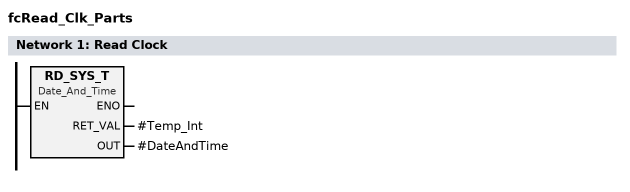
   #Temp_Int := RD_SYS_T(out => #DateAndTime);
END_REGION

REGION Network 2 (STL)

         LAR1  #""Address_4";
         L     B[AR1, P#0.0];
         T     #Year;
         L     B[AR1, P#1.0];
         T     #Month;
         L     B[AR1, P#2.0];
         T     #Day;
         L     B[AR1, P#3.0];
         T     #Hour;
         L     B[AR1, P#4.0];
         T     #Minute;
         L     B[AR1, P#5.0];
         T     #Second;

         L     W#16#FFF0;
         L     W[AR1, P#6.0];
         AW;
         T     #MilliSecond;

         L     B#16#F;
         L     B[AR1, P#7.0];
         AW;
         T     #DayOfWeek;
         CLR;
END_REGION
END_FUNCTION

FUNCTION "fcByteToBits" : Void   // FC1002, LAD
TITLE = Split byte into bits
{ S7_Optimized_Access := 'FALSE' }
VERSION : 0.1
BEGIN

REGION Network 1: Bit 0
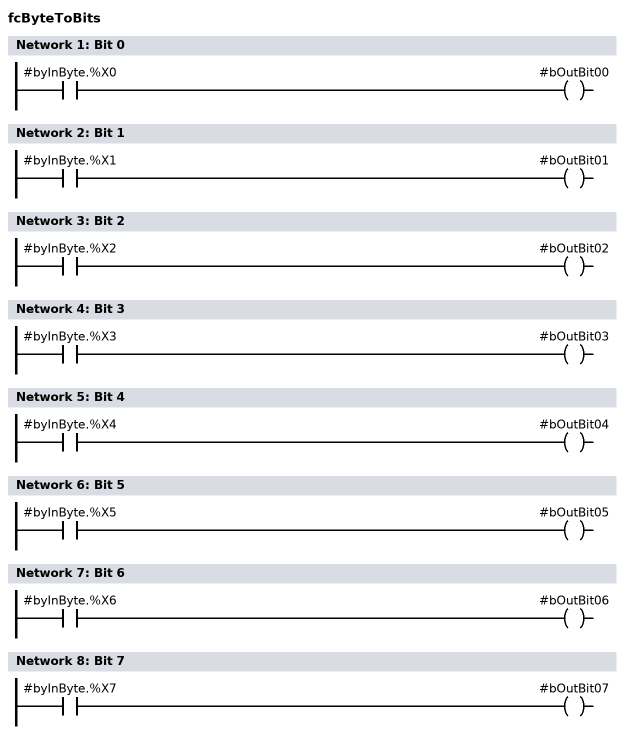
   RUNG wire#powerrail
      Contact( #byInByte.%X0 )
      Coil( #bOutBit00 )
   END_RUNG
   // the same network as SCL:
   #bOutBit00 := #byInByte.%X0;
END_REGION

REGION Network 2: Bit 1
   RUNG wire#powerrail
      Contact( #byInByte.%X1 )
      Coil( #bOutBit01 )
   END_RUNG
   // the same network as SCL:
   #bOutBit01 := #byInByte.%X1;
END_REGION

REGION Network 3: Bit 2
   RUNG wire#powerrail
      Contact( #byInByte.%X2 )
      Coil( #bOutBit02 )
   END_RUNG
   // the same network as SCL:
   #bOutBit02 := #byInByte.%X2;
END_REGION

REGION Network 4: Bit 3
   RUNG wire#powerrail
      Contact( #byInByte.%X3 )
      Coil( #bOutBit03 )
   END_RUNG
   // the same network as SCL:
   #bOutBit03 := #byInByte.%X3;
END_REGION

REGION Network 5: Bit 4
   RUNG wire#powerrail
      Contact( #byInByte.%X4 )
      Coil( #bOutBit04 )
   END_RUNG
   // the same network as SCL:
   #bOutBit04 := #byInByte.%X4;
END_REGION

REGION Network 6: Bit 5
   RUNG wire#powerrail
      Contact( #byInByte.%X5 )
      Coil( #bOutBit05 )
   END_RUNG
   // the same network as SCL:
   #bOutBit05 := #byInByte.%X5;
END_REGION

REGION Network 7: Bit 6
   RUNG wire#powerrail
      Contact( #byInByte.%X6 )
      Coil( #bOutBit06 )
   END_RUNG
   // the same network as SCL:
   #bOutBit06 := #byInByte.%X6;
END_REGION

REGION Network 8: Bit 7
   RUNG wire#powerrail
      Contact( #byInByte.%X7 )
      Coil( #bOutBit07 )
   END_RUNG
   // the same network as SCL:
   #bOutBit07 := #byInByte.%X7;
END_REGION
END_FUNCTION

FUNCTION "fbBitsToByte" : Void   // FC1003, LAD
TITLE = Pack bits into byte
{ S7_Optimized_Access := 'FALSE' }
VERSION : 0.1
BEGIN

REGION Network 1: Bit0
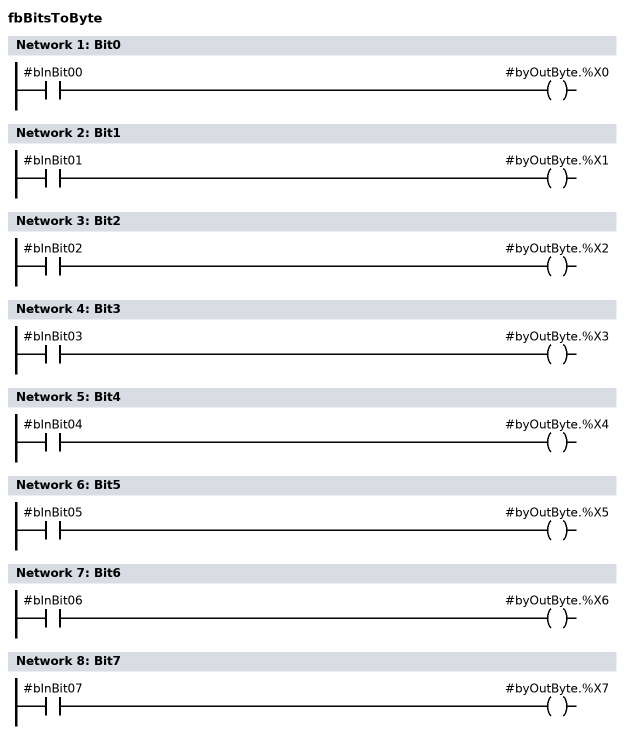
   RUNG wire#powerrail
      Contact( #bInBit00 )
      Coil( #byOutByte.%X0 )
   END_RUNG
   // the same network as SCL:
   #byOutByte.%X0 := #bInBit00;
END_REGION

REGION Network 2: Bit1
   RUNG wire#powerrail
      Contact( #bInBit01 )
      Coil( #byOutByte.%X1 )
   END_RUNG
   // the same network as SCL:
   #byOutByte.%X1 := #bInBit01;
END_REGION

REGION Network 3: Bit2
   RUNG wire#powerrail
      Contact( #bInBit02 )
      Coil( #byOutByte.%X2 )
   END_RUNG
   // the same network as SCL:
   #byOutByte.%X2 := #bInBit02;
END_REGION

REGION Network 4: Bit3
   RUNG wire#powerrail
      Contact( #bInBit03 )
      Coil( #byOutByte.%X3 )
   END_RUNG
   // the same network as SCL:
   #byOutByte.%X3 := #bInBit03;
END_REGION

REGION Network 5: Bit4
   RUNG wire#powerrail
      Contact( #bInBit04 )
      Coil( #byOutByte.%X4 )
   END_RUNG
   // the same network as SCL:
   #byOutByte.%X4 := #bInBit04;
END_REGION

REGION Network 6: Bit5
   RUNG wire#powerrail
      Contact( #bInBit05 )
      Coil( #byOutByte.%X5 )
   END_RUNG
   // the same network as SCL:
   #byOutByte.%X5 := #bInBit05;
END_REGION

REGION Network 7: Bit6
   RUNG wire#powerrail
      Contact( #bInBit06 )
      Coil( #byOutByte.%X6 )
   END_RUNG
   // the same network as SCL:
   #byOutByte.%X6 := #bInBit06;
END_REGION

REGION Network 8: Bit7
   RUNG wire#powerrail
      Contact( #bInBit07 )
      Coil( #byOutByte.%X7 )
   END_RUNG
   // the same network as SCL:
   #byOutByte.%X7 := #bInBit07;
END_REGION
END_FUNCTION

FUNCTION "fcCreateAnyPointer" : Void   // FC1025, STL
TITLE = Creates any pointer
{ S7_Optimized_Access := 'FALSE' }
VERSION : 0.1
BEGIN

REGION Network 1: It won't work in LAD, STL only
   // Create pointer in the temp location (AR1)
         LAR1  #""Address_2";

   // Syntax ID - always 10
         L     B#16#10;
         T     LB[AR1, P#0.0];

   // Data type
         L     #byInDataType;
         T     LB[AR1, P#1.0];

   // Size
         L     #iInSize;
         T     LW[AR1, P#2.0];

   // DB number
         L     #iInDB_Num;
         T     LW[AR1, P#4.0];


   // Memory area
         L     #byInMemoryArea;
         T     LB[AR1, P#6.0];

   // Offset high byte
         L     #iInOffsetByte;
         SRD   13;
         T     LB[AR1, P#7.0];

   // Offset low word
         L     #iInOffsetBit;
         AW    16#0007;

         L     #iInOffsetByte;
         SLD   3;

         OW;
         T     LW[AR1, P#8.0];

   // Write to the output (AR2)
         L     #""Address_21";
         LAR2;

         L     LD[AR1, P#0.0];
         T     D[AR2, P#0.0];

         L     LD[AR1, P#4.0];
         T     D[AR2, P#4.0];

         L     LW[AR1, P#8.0];
         T     W[AR2, P#8.0];
END_REGION

REGION Network 2
         SET;
         SAVE;
END_REGION
END_FUNCTION

FUNCTION "fcParseAnyPointer" : Void   // FC1026, SCL
{ S7_Optimized_Access := 'FALSE' }
VERSION : 0.0
BEGIN


       #AnyPointer := #pInAnyPointer;

       #AnyStruc.SyntaxID := b#16#10;
       #byOutDataType := #AnyStruc.DataType;
       #iOutSize := WORD_TO_INT(#AnyStruc.Size);
       #iOutDB_Num := WORD_TO_INT(#AnyStruc.DB_Num);
       #byOutMemoryArea := #AnyStruc.MemoryArea;
       #iOutOffsetBit := WORD_TO_INT(#AnyStruc.OffsetLo AND w#16#0007);
       #iOutOffsetByte := WORD_TO_INT(SHR(IN := #AnyStruc.OffsetLo, N := 3) OR SHL(IN := BYTE_TO_WORD(#AnyStruc.OffsetHi), N := 13));

       ENO:=true;
END_FUNCTION

FUNCTION "fcTemperatureConvert" : Void   // FC1027, LAD
{ S7_Optimized_Access := 'FALSE' }
VERSION : 0.1
BEGIN

REGION Network 1: Convert F to C
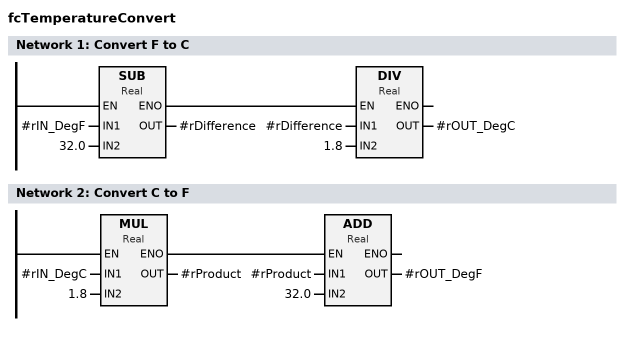
   RUNG wire#powerrail
      { S7_Templates := "SrcType := Real"; S7_GenerateENO := "TRUE" } Sub(in1 := #rIN_DegF, in2 := 32.0, out => #rDifference)
      { S7_Templates := "SrcType := Real"; S7_GenerateENO := "TRUE" } Div(in1 := #rDifference, in2 := 1.8, out => #rOUT_DegC)
   END_RUNG
   // the same network as SCL:
   // ENO of a box is taken as its EN; it also drops when the box reports an error
   #rDifference := #rIN_DegF - 32.0;
   #rOUT_DegC := #rDifference / 1.8;
END_REGION

REGION Network 2: Convert C to F
   RUNG wire#powerrail
      { S7_Templates := "SrcType := Real"; S7_GenerateENO := "TRUE" } Mul(in1 := #rIN_DegC, in2 := 1.8, out => #rProduct)
      { S7_Templates := "SrcType := Real"; S7_GenerateENO := "TRUE" } Add(in1 := #rProduct, in2 := 32.0, out => #rOUT_DegF)
   END_RUNG
   // the same network as SCL:
   // ENO of a box is taken as its EN; it also drops when the box reports an error
   #rProduct := #rIN_DegC * 1.8;
   #rOUT_DegF := #rProduct + 32.0;
END_REGION
END_FUNCTION

// folder: Resources/IO

FUNCTION "fcReadInput_LinearScale" : Void   // FC308, LAD
TITLE = Read/Scale input word
{ S7_Optimized_Access := 'FALSE' }
VERSION : 0.1
BEGIN

REGION Network 1: Swap input value bytes if needed
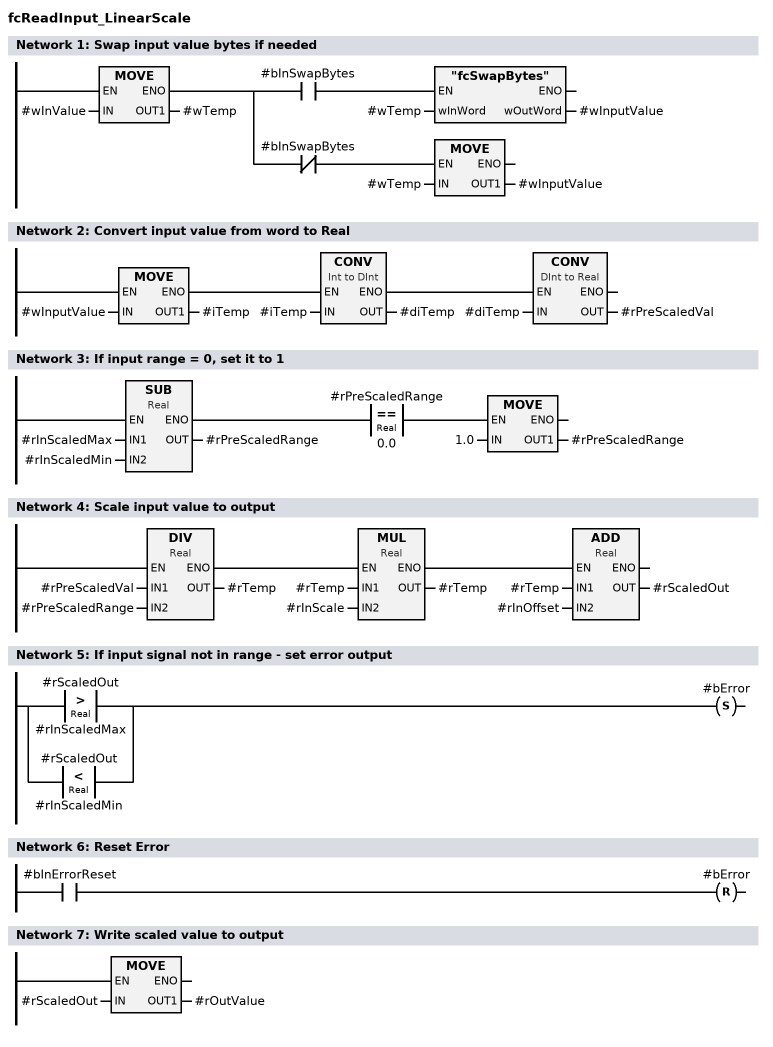
   RUNG wire#powerrail
      { S7_GenerateENO := "TRUE" } Move(in := #wInValue, out1 => #wTemp)
      wire#w1
      Contact( #bInSwapBytes )
      "fcSwapBytes"(wInWord := #wTemp, wOutWord => #wInputValue)
   END_RUNG
   RUNG wire#w1
      I_Contact( #bInSwapBytes )
      { S7_GenerateENO := "TRUE" } Move(in := #wTemp, out1 => #wInputValue)
   END_RUNG
   // the same network as SCL:
   // ENO of a box is taken as its EN; it also drops when the box reports an error
   #wTemp := #wInValue;
   IF #bInSwapBytes THEN "fcSwapBytes"(wInWord := #wTemp, wOutWord => #wInputValue); END_IF;
   IF NOT #bInSwapBytes THEN #wInputValue := #wTemp; END_IF;
END_REGION

REGION Network 2: Convert input value from word to Real
   RUNG wire#powerrail
      { S7_GenerateENO := "TRUE" } Move(in := #wInputValue, out1 => #iTemp)
      { S7_Templates := "[SrcType := Int, DestType := DInt]"; S7_GenerateENO := "TRUE" } Convert(in := #iTemp, out => #diTemp)
      { S7_Templates := "[SrcType := DInt, DestType := Real]"; S7_GenerateENO := "TRUE" } Convert(in := #diTemp, out => #rPreScaledVal)
   END_RUNG
   // the same network as SCL:
   // ENO of a box is taken as its EN; it also drops when the box reports an error
   #iTemp := #wInputValue;
   #diTemp := INT_TO_DINT(#iTemp);
   #rPreScaledVal := DINT_TO_REAL(#diTemp);
END_REGION

REGION Network 3: If input range = 0, set it to 1
   RUNG wire#powerrail
      { S7_Templates := "SrcType := Real"; S7_GenerateENO := "TRUE" } Sub(in1 := #rInScaledMax, in2 := #rInScaledMin, out => #rPreScaledRange)
      { S7_Templates := "SrcType := Real" } EQ_Contact(in1 := #rPreScaledRange, in2 := 0.0)
      { S7_GenerateENO := "TRUE" } Move(in := 1.0, out1 => #rPreScaledRange)
   END_RUNG
   // the same network as SCL:
   // ENO of a box is taken as its EN; it also drops when the box reports an error
   #rPreScaledRange := #rInScaledMax - #rInScaledMin;
   IF #rPreScaledRange = 0.0 THEN #rPreScaledRange := 1.0; END_IF;
END_REGION

REGION Network 4: Scale input value to output
   RUNG wire#powerrail
      { S7_Templates := "SrcType := Real"; S7_GenerateENO := "TRUE" } Div(in1 := #rPreScaledVal, in2 := #rPreScaledRange, out => #rTemp)
      { S7_Templates := "SrcType := Real"; S7_GenerateENO := "TRUE" } Mul(in1 := #rTemp, in2 := #rInScale, out => #rTemp)
      { S7_Templates := "SrcType := Real"; S7_GenerateENO := "TRUE" } Add(in1 := #rTemp, in2 := #rInOffset, out => #rScaledOut)
   END_RUNG
   // the same network as SCL:
   // ENO of a box is taken as its EN; it also drops when the box reports an error
   #rTemp := #rPreScaledVal / #rPreScaledRange;
   #rTemp := #rTemp * #rInScale;
   #rScaledOut := #rTemp + #rInOffset;
END_REGION

REGION Network 5: If input signal not in range - set error output
   RUNG wire#powerrail
      { S7_Templates := "SrcType := Real" } GT_Contact(in1 := #rScaledOut, in2 := #rInScaledMax)
      wire#w1
      S_Coil( #bError )
   END_RUNG
   RUNG wire#powerrail
      { S7_Templates := "SrcType := Real" } LT_Contact(in1 := #rScaledOut, in2 := #rInScaledMin)
   END_RUNG wire#w1
   // the same network as SCL:
   IF (#rScaledOut > #rInScaledMax) OR (#rScaledOut < #rInScaledMin) THEN #bError := TRUE; END_IF;
END_REGION

REGION Network 6: Reset Error
   RUNG wire#powerrail
      Contact( #bInErrorReset )
      R_Coil( #bError )
   END_RUNG
   // the same network as SCL:
   IF #bInErrorReset THEN #bError := FALSE; END_IF;
END_REGION

REGION Network 7: Write scaled value to output
   RUNG wire#powerrail
      { S7_GenerateENO := "TRUE" } Move(in := #rScaledOut, out1 => #rOutValue)
   END_RUNG
   // the same network as SCL:
   #rOutValue := #rScaledOut;
END_REGION

REGION Network 8 (STL): Set ENO
         SET;
         SAVE;
END_REGION
END_FUNCTION

FUNCTION "fcReadInput_LinearScale" : Void   // FC308, LAD
TITLE = Read/Scale input word
{ S7_Optimized_Access := 'FALSE' }
VERSION : 0.1
BEGIN

REGION Network 1: Swap input value bytes if needed
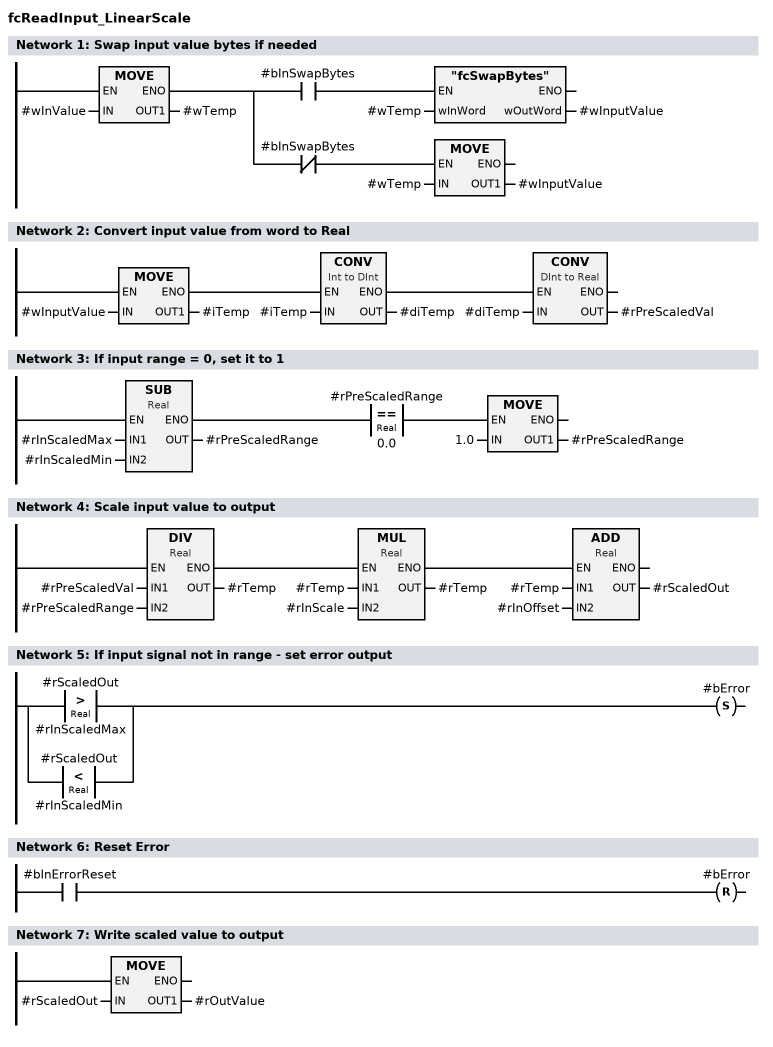
   RUNG wire#powerrail
      { S7_GenerateENO := "TRUE" } Move(in := #wInValue, out1 => #wTemp)
      wire#w1
      Contact( #bInSwapBytes )
      "fcSwapBytes"(wInWord := #wTemp, wOutWord => #wInputValue)
   END_RUNG
   RUNG wire#w1
      I_Contact( #bInSwapBytes )
      { S7_GenerateENO := "TRUE" } Move(in := #wTemp, out1 => #wInputValue)
   END_RUNG
   // the same network as SCL:
   // ENO of a box is taken as its EN; it also drops when the box reports an error
   #wTemp := #wInValue;
   IF #bInSwapBytes THEN "fcSwapBytes"(wInWord := #wTemp, wOutWord => #wInputValue); END_IF;
   IF NOT #bInSwapBytes THEN #wInputValue := #wTemp; END_IF;
END_REGION

REGION Network 2: Convert input value from word to Real
   RUNG wire#powerrail
      { S7_GenerateENO := "TRUE" } Move(in := #wInputValue, out1 => #iTemp)
      { S7_Templates := "[SrcType := Int, DestType := DInt]"; S7_GenerateENO := "TRUE" } Convert(in := #iTemp, out => #diTemp)
      { S7_Templates := "[SrcType := DInt, DestType := Real]"; S7_GenerateENO := "TRUE" } Convert(in := #diTemp, out => #rPreScaledVal)
   END_RUNG
   // the same network as SCL:
   // ENO of a box is taken as its EN; it also drops when the box reports an error
   #iTemp := #wInputValue;
   #diTemp := INT_TO_DINT(#iTemp);
   #rPreScaledVal := DINT_TO_REAL(#diTemp);
END_REGION

REGION Network 3: If input range = 0, set it to 1
   RUNG wire#powerrail
      { S7_Templates := "SrcType := Real"; S7_GenerateENO := "TRUE" } Sub(in1 := #rInScaledMax, in2 := #rInScaledMin, out => #rPreScaledRange)
      { S7_Templates := "SrcType := Real" } EQ_Contact(in1 := #rPreScaledRange, in2 := 0.0)
      { S7_GenerateENO := "TRUE" } Move(in := 1.0, out1 => #rPreScaledRange)
   END_RUNG
   // the same network as SCL:
   // ENO of a box is taken as its EN; it also drops when the box reports an error
   #rPreScaledRange := #rInScaledMax - #rInScaledMin;
   IF #rPreScaledRange = 0.0 THEN #rPreScaledRange := 1.0; END_IF;
END_REGION

REGION Network 4: Scale input value to output
   RUNG wire#powerrail
      { S7_Templates := "SrcType := Real"; S7_GenerateENO := "TRUE" } Div(in1 := #rPreScaledVal, in2 := #rPreScaledRange, out => #rTemp)
      { S7_Templates := "SrcType := Real"; S7_GenerateENO := "TRUE" } Mul(in1 := #rTemp, in2 := #rInScale, out => #rTemp)
      { S7_Templates := "SrcType := Real"; S7_GenerateENO := "TRUE" } Add(in1 := #rTemp, in2 := #rInOffset, out => #rScaledOut)
   END_RUNG
   // the same network as SCL:
   // ENO of a box is taken as its EN; it also drops when the box reports an error
   #rTemp := #rPreScaledVal / #rPreScaledRange;
   #rTemp := #rTemp * #rInScale;
   #rScaledOut := #rTemp + #rInOffset;
END_REGION

REGION Network 5: If input signal not in range - set error output
   RUNG wire#powerrail
      { S7_Templates := "SrcType := Real" } GT_Contact(in1 := #rScaledOut, in2 := #rInScaledMax)
      wire#w1
      S_Coil( #bError )
   END_RUNG
   RUNG wire#powerrail
      { S7_Templates := "SrcType := Real" } LT_Contact(in1 := #rScaledOut, in2 := #rInScaledMin)
   END_RUNG wire#w1
   // the same network as SCL:
   IF (#rScaledOut > #rInScaledMax) OR (#rScaledOut < #rInScaledMin) THEN #bError := TRUE; END_IF;
END_REGION

REGION Network 6: Reset Error
   RUNG wire#powerrail
      Contact( #bInErrorReset )
      R_Coil( #bError )
   END_RUNG
   // the same network as SCL:
   IF #bInErrorReset THEN #bError := FALSE; END_IF;
END_REGION

REGION Network 7: Write scaled value to output
   RUNG wire#powerrail
      { S7_GenerateENO := "TRUE" } Move(in := #rScaledOut, out1 => #rOutValue)
   END_RUNG
   // the same network as SCL:
   #rOutValue := #rScaledOut;
END_REGION
END_FUNCTION

FUNCTION "fcWriteOutput_LinearScale" : Void   // FC309, LAD
TITLE = Scales an input to a specified slope and offset
{ S7_Optimized_Access := 'FALSE' }
VERSION : 0.1
BEGIN

REGION Network 1: Calculate total range of scale
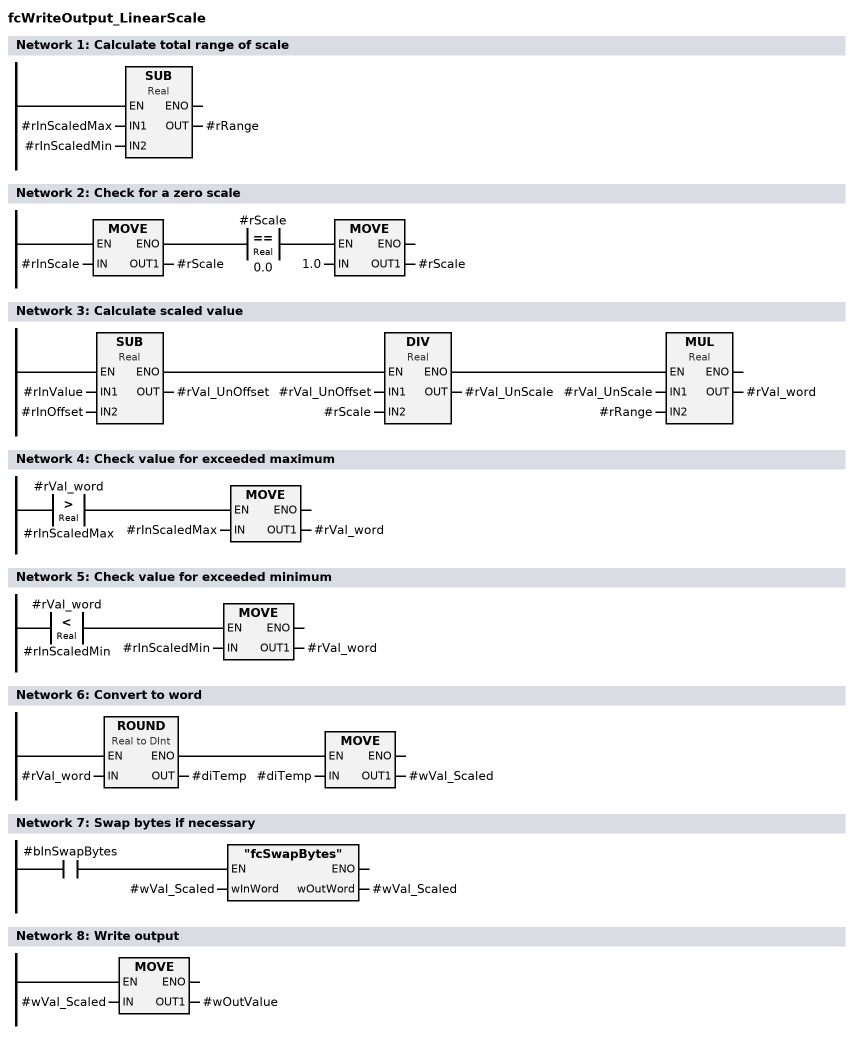
   RUNG wire#powerrail
      { S7_Templates := "SrcType := Real"; S7_GenerateENO := "TRUE" } Sub(in1 := #rInScaledMax, in2 := #rInScaledMin, out => #rRange)
   END_RUNG
   // the same network as SCL:
   #rRange := #rInScaledMax - #rInScaledMin;
END_REGION

REGION Network 2: Check for a zero scale
   RUNG wire#powerrail
      { S7_GenerateENO := "TRUE" } Move(in := #rInScale, out1 => #rScale)
      { S7_Templates := "SrcType := Real" } EQ_Contact(in1 := #rScale, in2 := 0.0)
      { S7_GenerateENO := "TRUE" } Move(in := 1.0, out1 => #rScale)
   END_RUNG
   // the same network as SCL:
   // ENO of a box is taken as its EN; it also drops when the box reports an error
   #rScale := #rInScale;
   IF #rScale = 0.0 THEN #rScale := 1.0; END_IF;
END_REGION

REGION Network 3: Calculate scaled value
   RUNG wire#powerrail
      { S7_Templates := "SrcType := Real"; S7_GenerateENO := "TRUE" } Sub(in1 := #rInValue, in2 := #rInOffset, out => #rVal_UnOffset)
      { S7_Templates := "SrcType := Real"; S7_GenerateENO := "TRUE" } Div(in1 := #rVal_UnOffset, in2 := #rScale, out => #rVal_UnScale)
      { S7_Templates := "SrcType := Real"; S7_GenerateENO := "TRUE" } Mul(in1 := #rVal_UnScale, in2 := #rRange, out => #rVal_word)
   END_RUNG
   // the same network as SCL:
   // ENO of a box is taken as its EN; it also drops when the box reports an error
   #rVal_UnOffset := #rInValue - #rInOffset;
   #rVal_UnScale := #rVal_UnOffset / #rScale;
   #rVal_word := #rVal_UnScale * #rRange;
END_REGION

REGION Network 4: Check value for exceeded maximum
   RUNG wire#powerrail
      { S7_Templates := "SrcType := Real" } GT_Contact(in1 := #rVal_word, in2 := #rInScaledMax)
      { S7_GenerateENO := "TRUE" } Move(in := #rInScaledMax, out1 => #rVal_word)
   END_RUNG
   // the same network as SCL:
   IF #rVal_word > #rInScaledMax THEN #rVal_word := #rInScaledMax; END_IF;
END_REGION

REGION Network 5: Check value for exceeded minimum
   RUNG wire#powerrail
      { S7_Templates := "SrcType := Real" } LT_Contact(in1 := #rVal_word, in2 := #rInScaledMin)
      { S7_GenerateENO := "TRUE" } Move(in := #rInScaledMin, out1 => #rVal_word)
   END_RUNG
   // the same network as SCL:
   IF #rVal_word < #rInScaledMin THEN #rVal_word := #rInScaledMin; END_IF;
END_REGION

REGION Network 6: Convert to word
   RUNG wire#powerrail
      { S7_Templates := "[SrcType := Real, DestType := DInt]"; S7_GenerateENO := "TRUE" } Round(in := #rVal_word, out => #diTemp)
      { S7_GenerateENO := "TRUE" } Move(in := #diTemp, out1 => #wVal_Scaled)
   END_RUNG
   // the same network as SCL:
   // ENO of a box is taken as its EN; it also drops when the box reports an error
   #diTemp := ROUND(#rVal_word);
   #wVal_Scaled := #diTemp;
END_REGION

REGION Network 7: Swap bytes if necessary
   RUNG wire#powerrail
      Contact( #bInSwapBytes )
      "fcSwapBytes"(wInWord := #wVal_Scaled, wOutWord => #wVal_Scaled)
   END_RUNG
   // the same network as SCL:
   IF #bInSwapBytes THEN "fcSwapBytes"(wInWord := #wVal_Scaled, wOutWord => #wVal_Scaled); END_IF;
END_REGION

REGION Network 8: Write output
   RUNG wire#powerrail
      { S7_GenerateENO := "TRUE" } Move(in := #wVal_Scaled, out1 => #wOutValue)
   END_RUNG
   // the same network as SCL:
   #wOutValue := #wVal_Scaled;
END_REGION

REGION Network 9 (STL): Set RLO
         SET;
         SAVE;
END_REGION
END_FUNCTION

FUNCTION "fcWriteOutput_LinearScale" : Void   // FC309, LAD
TITLE = Scales an input to a specified slope and offset
{ S7_Optimized_Access := 'FALSE' }
VERSION : 0.1
BEGIN

REGION Network 1: Calculate total range of scale
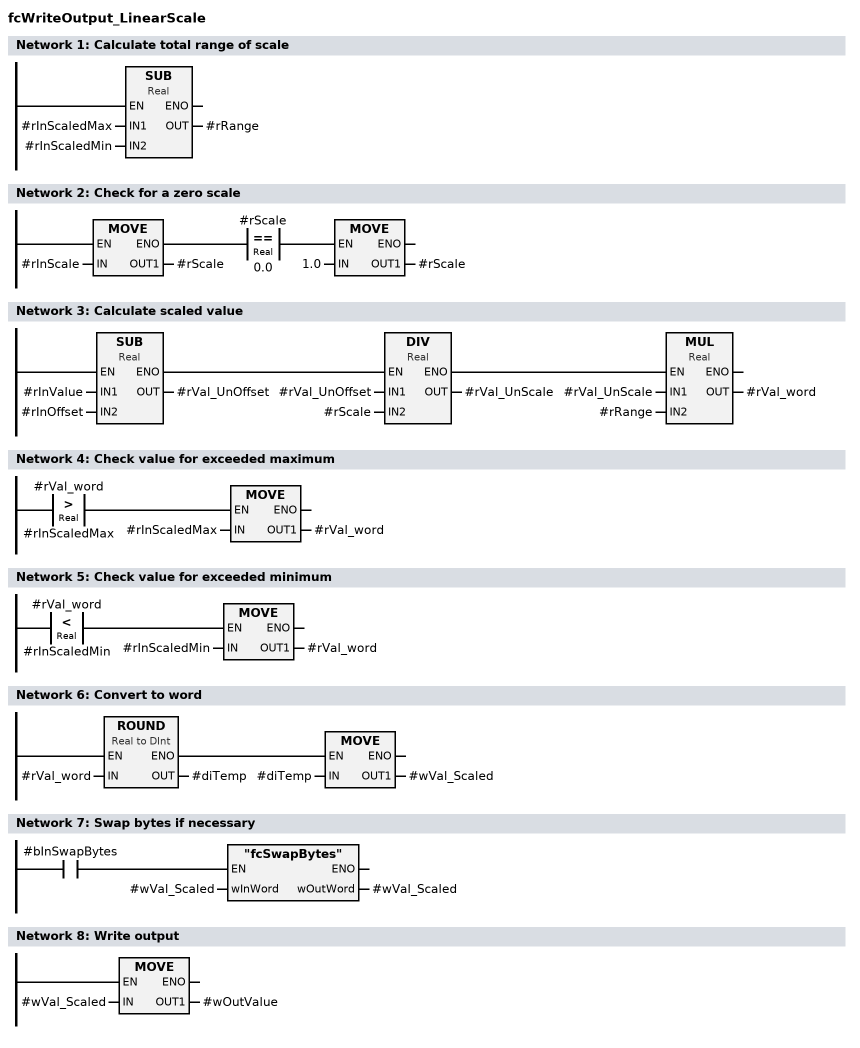
   RUNG wire#powerrail
      { S7_Templates := "SrcType := Real"; S7_GenerateENO := "TRUE" } Sub(in1 := #rInScaledMax, in2 := #rInScaledMin, out => #rRange)
   END_RUNG
   // the same network as SCL:
   #rRange := #rInScaledMax - #rInScaledMin;
END_REGION

REGION Network 2: Check for a zero scale
   RUNG wire#powerrail
      { S7_GenerateENO := "TRUE" } Move(in := #rInScale, out1 => #rScale)
      { S7_Templates := "SrcType := Real" } EQ_Contact(in1 := #rScale, in2 := 0.0)
      { S7_GenerateENO := "TRUE" } Move(in := 1.0, out1 => #rScale)
   END_RUNG
   // the same network as SCL:
   // ENO of a box is taken as its EN; it also drops when the box reports an error
   #rScale := #rInScale;
   IF #rScale = 0.0 THEN #rScale := 1.0; END_IF;
END_REGION

REGION Network 3: Calculate scaled value
   RUNG wire#powerrail
      { S7_Templates := "SrcType := Real"; S7_GenerateENO := "TRUE" } Sub(in1 := #rInValue, in2 := #rInOffset, out => #rVal_UnOffset)
      { S7_Templates := "SrcType := Real"; S7_GenerateENO := "TRUE" } Div(in1 := #rVal_UnOffset, in2 := #rScale, out => #rVal_UnScale)
      { S7_Templates := "SrcType := Real"; S7_GenerateENO := "TRUE" } Mul(in1 := #rVal_UnScale, in2 := #rRange, out => #rVal_word)
   END_RUNG
   // the same network as SCL:
   // ENO of a box is taken as its EN; it also drops when the box reports an error
   #rVal_UnOffset := #rInValue - #rInOffset;
   #rVal_UnScale := #rVal_UnOffset / #rScale;
   #rVal_word := #rVal_UnScale * #rRange;
END_REGION

REGION Network 4: Check value for exceeded maximum
   RUNG wire#powerrail
      { S7_Templates := "SrcType := Real" } GT_Contact(in1 := #rVal_word, in2 := #rInScaledMax)
      { S7_GenerateENO := "TRUE" } Move(in := #rInScaledMax, out1 => #rVal_word)
   END_RUNG
   // the same network as SCL:
   IF #rVal_word > #rInScaledMax THEN #rVal_word := #rInScaledMax; END_IF;
END_REGION

REGION Network 5: Check value for exceeded minimum
   RUNG wire#powerrail
      { S7_Templates := "SrcType := Real" } LT_Contact(in1 := #rVal_word, in2 := #rInScaledMin)
      { S7_GenerateENO := "TRUE" } Move(in := #rInScaledMin, out1 => #rVal_word)
   END_RUNG
   // the same network as SCL:
   IF #rVal_word < #rInScaledMin THEN #rVal_word := #rInScaledMin; END_IF;
END_REGION

REGION Network 6: Convert to word
   RUNG wire#powerrail
      { S7_Templates := "[SrcType := Real, DestType := DInt]"; S7_GenerateENO := "TRUE" } Round(in := #rVal_word, out => #diTemp)
      { S7_GenerateENO := "TRUE" } Move(in := #diTemp, out1 => #wVal_Scaled)
   END_RUNG
   // the same network as SCL:
   // ENO of a box is taken as its EN; it also drops when the box reports an error
   #diTemp := ROUND(#rVal_word);
   #wVal_Scaled := #diTemp;
END_REGION

REGION Network 7: Swap bytes if necessary
   RUNG wire#powerrail
      Contact( #bInSwapBytes )
      "fcSwapBytes"(wInWord := #wVal_Scaled, wOutWord => #wVal_Scaled)
   END_RUNG
   // the same network as SCL:
   IF #bInSwapBytes THEN "fcSwapBytes"(wInWord := #wVal_Scaled, wOutWord => #wVal_Scaled); END_IF;
END_REGION

REGION Network 8: Write output
   RUNG wire#powerrail
      { S7_GenerateENO := "TRUE" } Move(in := #wVal_Scaled, out1 => #wOutValue)
   END_RUNG
   // the same network as SCL:
   #wOutValue := #wVal_Scaled;
END_REGION
END_FUNCTION

FUNCTION "fcReadPID" : Void   // FC1037, SCL
TITLE = fcReadPID
{ S7_Optimized_Access := 'FALSE' }
AUTHOR : DMC
FAMILY : IO
NAME : RD_PID
VERSION : 1.0
// This block read a peripheral input word
//  To use this block, feed in the address of the PID you would like to read
//  for example: to read PID123 you would input the number 123 to the input iPID_Address
//  the entire word is read and output as wPID_Value
//  Block Parameters
BEGIN


   //this reads the word from the specified peripheral input
   #dwOutValue:=%ID(#iInAddress):P;

   ENO:=TRUE;
END_FUNCTION

FUNCTION "fcReadPID" : Void   // FC1037, SCL
TITLE = fcReadPID
{ S7_Optimized_Access := 'FALSE' }
AUTHOR : DMC
FAMILY : IO
NAME : RD_PID
VERSION : 1.0
// This block read a peripheral input word
//  To use this block, feed in the address of the PID you would like to read
//  for example: to read PID123 you would input the number 123 to the input iPID_Address
//  the entire word is read and output as wPID_Value
//  Block Parameters
BEGIN


   //this reads the word from the specified peripheral input
   #dwOutValue := PEEK(area := #cbyPeripheralInputArea, byteOffset := #iInAddress, dbNumber := 0);

   ENO:=TRUE;
END_FUNCTION

FUNCTION "fcWritePQD" : Void   // FC1038, SCL
TITLE = fcWritePQD
{ S7_Optimized_Access := 'FALSE' }
AUTHOR : DMC
FAMILY : IO
NAME : WR_PQD
VERSION : 1.0
// This block writes a peripheral output double word
//  to use this block, enter the address of the Peripheral word and the word value.
//  for example, to set the value of PQD123 to 500, you would set iPQD_Address=123, and wPQD_Value=500
//  Block Parameters
BEGIN


   //this writes the double word from the specified peripheral input
   %QD(#iInAddress):P:=#dwInValue;

   ENO:=TRUE;
END_FUNCTION

FUNCTION "fcWritePQD" : Void   // FC1038, SCL
TITLE = fcWritePQD
{ S7_Optimized_Access := 'FALSE' }
AUTHOR : DMC
FAMILY : IO
NAME : WR_PQD
VERSION : 1.0
// This block writes a peripheral output double word
//  to use this block, enter the address of the Peripheral word and the word value.
//  for example, to set the value of PQD123 to 500, you would set iPQD_Address=123, and wPQD_Value=500
//  Block Parameters
BEGIN


   //this writes the double word from the specified peripheral input
   POKE(area := #cbyPeripheralOutputArea,
        byteOffset := #iInAddress,
        dbNumber := 0,
        value := #dwInValue);

   ENO:=TRUE;
END_FUNCTION

FUNCTION "fcReadPIB" : Void   // FC1039, SCL
TITLE = fcReadPIB
{ S7_Optimized_Access := 'FALSE' }
AUTHOR : DMC
FAMILY : IO
NAME : RD_PIB
VERSION : 1.0
// This block read a peripheral input word
//  To use this block, feed in the address of the PIB you would like to read
//  for example: to read PIB123 you would input the number 123 to the input iPIB_Address
//  the entire byte is read and output as byPIB_Value
//  Block Parameters
BEGIN


   //this reads the word from the specified peripheral input
   #byOutValue:=%IB(#iInAddress):P;

   ENO:=TRUE;
END_FUNCTION

FUNCTION "fcReadPIB" : Void   // FC1039, SCL
TITLE = fcReadPIB
{ S7_Optimized_Access := 'FALSE' }
AUTHOR : DMC
FAMILY : IO
NAME : RD_PIB
VERSION : 1.0
// This block read a peripheral input word
//  To use this block, feed in the address of the PIB you would like to read
//  for example: to read PIB123 you would input the number 123 to the input iPIB_Address
//  the entire byte is read and output as byPIB_Value
//  Block Parameters
BEGIN


   //this reads the word from the specified peripheral input
   #byOutValue := PEEK(area := #cbyPeripheralInputArea, dbNumber := 0, byteOffset := #iInAddress);

   ENO:=TRUE;
END_FUNCTION

FUNCTION "fcWritePQB" : Void   // FC1040, SCL
TITLE = fcWritePQB
{ S7_Optimized_Access := 'FALSE' }
AUTHOR : DMC
FAMILY : IO
NAME : WR_PQB
VERSION : 1.0
// This block writes a peripheral output byte
//  to use this block, enter the address of the Peripheral byte and the byte value.
//  for example, to set the value of PQB123 to 500, you would set iPQB_Address=123, and wPQB_Value=500
//  Block Parameters
BEGIN


   //this writes the byte from the specified peripheral input
   %QB(#iInAddress):P:=#byInValue;

   ENO:=TRUE;
END_FUNCTION

FUNCTION "fcWritePQB" : Void   // FC1040, SCL
TITLE = fcWritePQB
{ S7_Optimized_Access := 'FALSE' }
AUTHOR : DMC
FAMILY : IO
NAME : WR_PQB
VERSION : 1.0
// This block writes a peripheral output byte
//  to use this block, enter the address of the Peripheral byte and the byte value.
//  for example, to set the value of PQB123 to 500, you would set iPQB_Address=123, and wPQB_Value=500
//  Block Parameters
BEGIN


   //this writes the byte from the specified peripheral input
   POKE(area := #cbyPeripheralOutputArea,
        byteOffset := #iInAddress,
        dbNumber := 0,
        value := #byInValue);

   ENO:=TRUE;
END_FUNCTION

// folder: Resources/Process

FUNCTION_BLOCK "fbPWM"   // FB94, LAD
TITLE = PWM Control
{ S7_Optimized_Access := 'FALSE' }
VERSION : 0.1
// Pulse Width Modulation
BEGIN

REGION Network 1: Reset Counter
   // Reset the counter if requested.
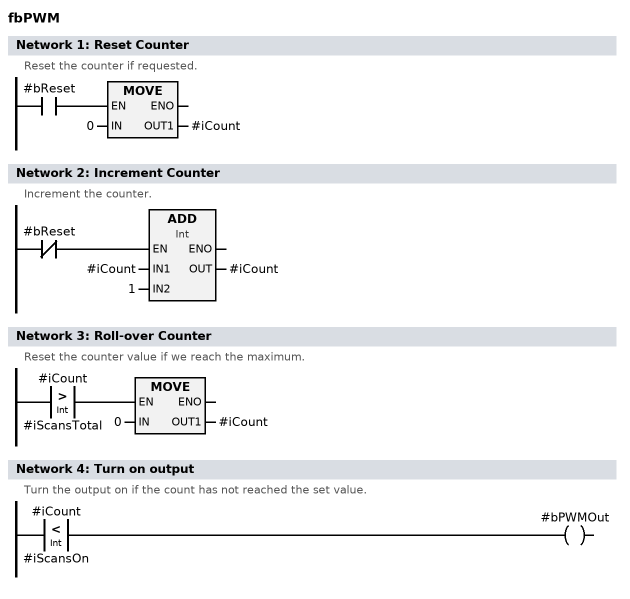
   RUNG wire#powerrail
      Contact( #bReset )
      { S7_GenerateENO := "TRUE" } Move(in := 0, out1 => #iCount)
   END_RUNG
   // the same network as SCL:
   IF #bReset THEN #iCount := 0; END_IF;
END_REGION

REGION Network 2: Increment Counter
   // Increment the counter.
   RUNG wire#powerrail
      I_Contact( #bReset )
      { S7_Templates := "SrcType := Int"; S7_GenerateENO := "TRUE" } Add(in1 := #iCount, in2 := 1, out => #iCount)
   END_RUNG
   // the same network as SCL:
   IF NOT #bReset THEN #iCount := #iCount + 1; END_IF;
END_REGION

REGION Network 3: Roll-over Counter
   // Reset the counter value if we reach the maximum.
   RUNG wire#powerrail
      { S7_Templates := "SrcType := Int" } GT_Contact(in1 := #iCount, in2 := #iScansTotal)
      { S7_GenerateENO := "TRUE" } Move(in := 0, out1 => #iCount)
   END_RUNG
   // the same network as SCL:
   IF #iCount > #iScansTotal THEN #iCount := 0; END_IF;
END_REGION

REGION Network 4: Turn on output
   // Turn the output on if the count has not reached the set value.
   RUNG wire#powerrail
      { S7_Templates := "SrcType := Int" } LT_Contact(in1 := #iCount, in2 := #iScansOn)
      Coil( #bPWMOut )
   END_RUNG
   // the same network as SCL:
   #bPWMOut := #iCount < #iScansOn;
END_REGION
END_FUNCTION_BLOCK

FUNCTION_BLOCK "fbPWMPhasedReset"   // FB95, LAD
TITLE = PWM Phased Reset Command
{ S7_Optimized_Access := 'FALSE' }
VERSION : 0.1
// Delays the PWM reset command a certain amount of scans based on this PWM's 
// index and total number of PWMs. Without this procedure, all of the PWMs would 
// turn on at the same time every period, causing a substantial, reoccuring 
// current 
// demand.
   VAR_TEMP   // added for the SCL form of the ladder/FBD networks
      _w1 : Bool;
      _w2 : Bool;
   END_VAR
BEGIN

REGION Network 1
   // Calculate the number of counts for this PWM object based on its index and total 
   // number of PWMs.